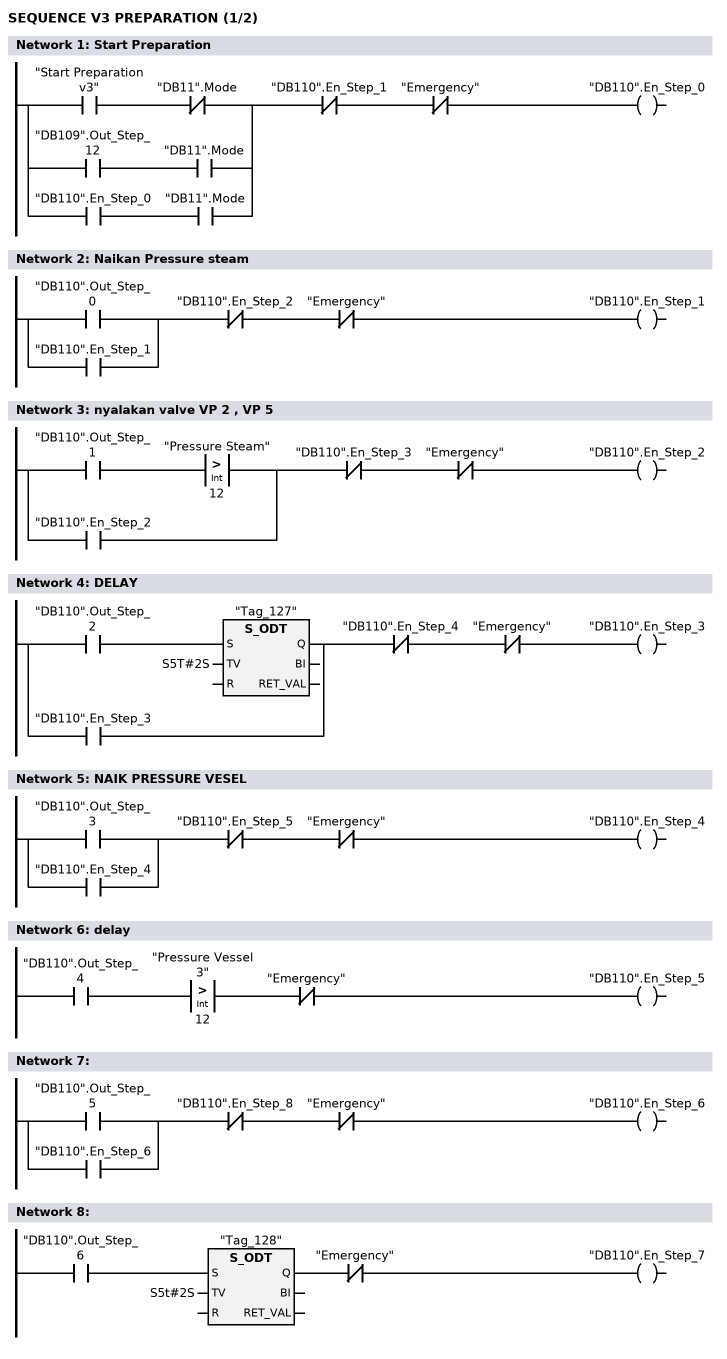
   RUNG wire#powerrail
      Contact( "Start Preparation v3" )
      I_Contact( "DB11".Mode )
      wire#w1
      I_Contact( "DB110".En_Step_1 )
      I_Contact( "Emergency" )
      Coil( "DB110".En_Step_0 )
   END_RUNG
   RUNG wire#powerrail
      Contact( "DB109".Out_Step_12 )
      Contact( "DB11".Mode )
   END_RUNG wire#w1
   RUNG wire#powerrail
      Contact( "DB110".En_Step_0 )
      Contact( "DB11".Mode )
   END_RUNG wire#w1
   // the same network as SCL:
   "DB110".En_Step_0 := (("Start Preparation v3" AND NOT "DB11".Mode) OR ("DB109".Out_Step_12 AND "DB11".Mode) OR ("DB110".En_Step_0 AND "DB11".Mode)) AND NOT "DB110".En_Step_1 AND NOT "Emergency";
END_REGION

REGION Network 2: Naikan Pressure steam
   RUNG wire#powerrail
      Contact( "DB110".Out_Step_0 )
      wire#w1
      I_Contact( "DB110".En_Step_2 )
      I_Contact( "Emergency" )
      Coil( "DB110".En_Step_1 )
   END_RUNG
   RUNG wire#powerrail
      Contact( "DB110".En_Step_1 )
   END_RUNG wire#w1
   // the same network as SCL:
   "DB110".En_Step_1 := ("DB110".Out_Step_0 OR "DB110".En_Step_1) AND NOT "DB110".En_Step_2 AND NOT "Emergency";
END_REGION

REGION Network 3: nyalakan valve VP 2 , VP 5
   RUNG wire#powerrail
      Contact( "DB110".Out_Step_1 )
      { S7_Templates := "SrcType := Int" } GT_Contact(in1 := "Pressure Steam", in2 := 12)
      wire#w1
      I_Contact( "DB110".En_Step_3 )
      I_Contact( "Emergency" )
      Coil( "DB110".En_Step_2 )
   END_RUNG
   RUNG wire#powerrail
      Contact( "DB110".En_Step_2 )
   END_RUNG wire#w1
   // the same network as SCL:
   "DB110".En_Step_2 := (("DB110".Out_Step_1 AND ("Pressure Steam" > 12)) OR "DB110".En_Step_2) AND NOT "DB110".En_Step_3 AND NOT "Emergency";
END_REGION

REGION Network 4: DELAY
   RUNG wire#powerrail
      Contact( "DB110".Out_Step_2 )
      S_ODT(T_NO := "Tag_127", TV := S5T#2S, R :=, BI =>, RET_VAL =>)
      wire#w1
      I_Contact( "DB110".En_Step_4 )
      I_Contact( "Emergency" )
      Coil( "DB110".En_Step_3 )
   END_RUNG
   RUNG wire#powerrail
      Contact( "DB110".En_Step_3 )
   END_RUNG wire#w1
   // the same network as SCL:
   #_s5time1 := S_ODT(T_NO := "Tag_127", S := "DB110".Out_Step_2, TV := S5T#2S, Q => #_w1);
   "DB110".En_Step_3 := (#_w1 OR "DB110".En_Step_3) AND NOT "DB110".En_Step_4 AND NOT "Emergency";
END_REGION

REGION Network 5: NAIK PRESSURE VESEL
   RUNG wire#powerrail
      Contact( "DB110".Out_Step_3 )
      wire#w1
      I_Contact( "DB110".En_Step_5 )
      I_Contact( "Emergency" )
      Coil( "DB110".En_Step_4 )
   END_RUNG
   RUNG wire#powerrail
      Contact( "DB110".En_Step_4 )
   END_RUNG wire#w1
   // the same network as SCL:
   "DB110".En_Step_4 := ("DB110".Out_Step_3 OR "DB110".En_Step_4) AND NOT "DB110".En_Step_5 AND NOT "Emergency";
END_REGION

REGION Network 6: delay
   RUNG wire#powerrail
      Contact( "DB110".Out_Step_4 )
      { S7_Templates := "SrcType := Int" } GT_Contact(in1 := "Pressure Vessel 3", in2 := 12)
      I_Contact( "Emergency" )
      Coil( "DB110".En_Step_5 )
   END_RUNG
   // the same network as SCL:
   "DB110".En_Step_5 := "DB110".Out_Step_4 AND ("Pressure Vessel 3" > 12) AND NOT "Emergency";
END_REGION

REGION Network 7
   RUNG wire#powerrail
      Contact( "DB110".Out_Step_5 )
      wire#w1
      I_Contact( "DB110".En_Step_8 )
      I_Contact( "Emergency" )
      Coil( "DB110".En_Step_6 )
   END_RUNG
   RUNG wire#powerrail
      Contact( "DB110".En_Step_6 )
   END_RUNG wire#w1
   // the same network as SCL:
   "DB110".En_Step_6 := ("DB110".Out_Step_5 OR "DB110".En_Step_6) AND NOT "DB110".En_Step_8 AND NOT "Emergency";
END_REGION

REGION Network 8
   RUNG wire#powerrail
      Contact( "DB110".Out_Step_6 )
      S_ODT(T_NO := "Tag_128", TV := S5t#2S, R :=, BI =>, RET_VAL =>)
      I_Contact( "Emergency" )
      Coil( "DB110".En_Step_7 )
   END_RUNG
   // the same network as SCL:
   #_s5time1 := S_ODT(T_NO := "Tag_128", S := "DB110".Out_Step_6, TV := S5t#2S, Q => #_w1);
   "DB110".En_Step_7 := #_w1 AND NOT "Emergency";
END_REGION

REGION Network 9: TURUNKAN PRESSURE
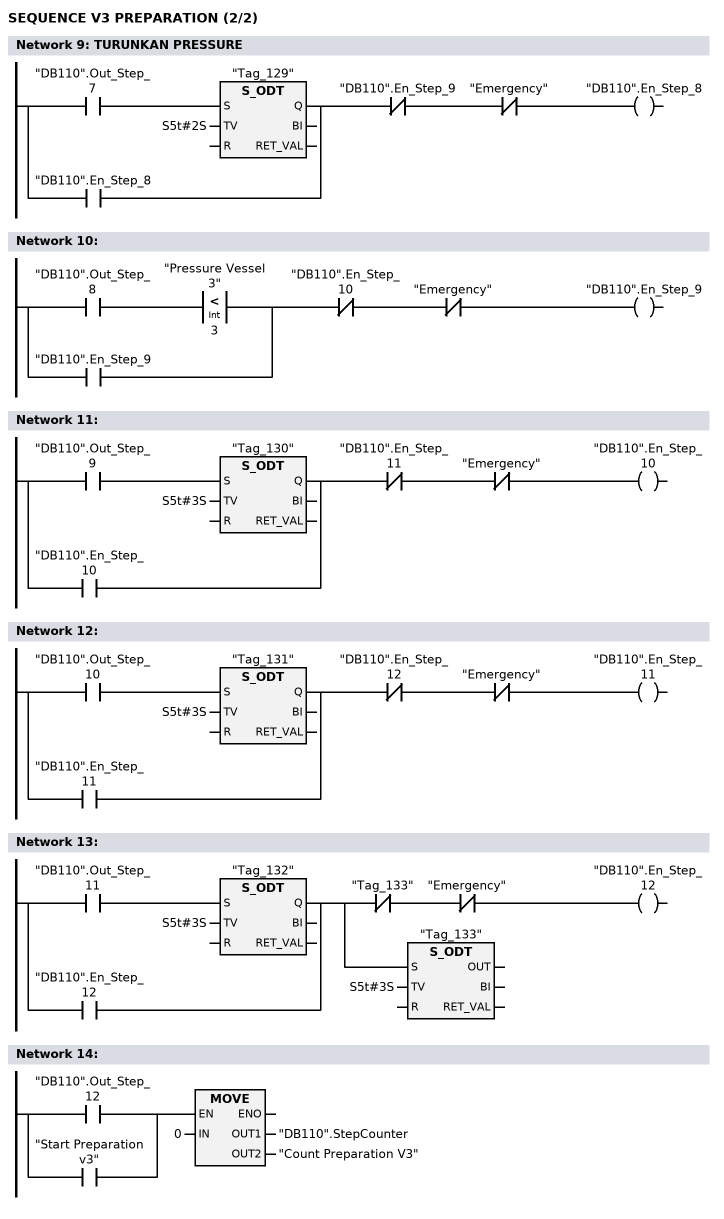
   RUNG wire#powerrail
      Contact( "DB110".Out_Step_7 )
      S_ODT(T_NO := "Tag_129", TV := S5t#2S, R :=, BI =>, RET_VAL =>)
      wire#w1
      I_Contact( "DB110".En_Step_9 )
      I_Contact( "Emergency" )
      Coil( "DB110".En_Step_8 )
   END_RUNG
   RUNG wire#powerrail
      Contact( "DB110".En_Step_8 )
   END_RUNG wire#w1
   // the same network as SCL:
   #_s5time1 := S_ODT(T_NO := "Tag_129", S := "DB110".Out_Step_7, TV := S5t#2S, Q => #_w1);
   "DB110".En_Step_8 := (#_w1 OR "DB110".En_Step_8) AND NOT "DB110".En_Step_9 AND NOT "Emergency";
END_REGION

REGION Network 10
   RUNG wire#powerrail
      Contact( "DB110".Out_Step_8 )
      { S7_Templates := "SrcType := Int" } LT_Contact(in1 := "Pressure Vessel 3", in2 := 3)
      wire#w1
      I_Contact( "DB110".En_Step_10 )
      I_Contact( "Emergency" )
      Coil( "DB110".En_Step_9 )
   END_RUNG
   RUNG wire#powerrail
      Contact( "DB110".En_Step_9 )
   END_RUNG wire#w1
   // the same network as SCL:
   "DB110".En_Step_9 := (("DB110".Out_Step_8 AND ("Pressure Vessel 3" < 3)) OR "DB110".En_Step_9) AND NOT "DB110".En_Step_10 AND NOT "Emergency";
END_REGION

REGION Network 11
   RUNG wire#powerrail
      Contact( "DB110".Out_Step_9 )
      S_ODT(T_NO := "Tag_130", TV := S5t#3S, R :=, BI =>, RET_VAL =>)
      wire#w1
      I_Contact( "DB110".En_Step_11 )
      I_Contact( "Emergency" )
      Coil( "DB110".En_Step_10 )
   END_RUNG
   RUNG wire#powerrail
      Contact( "DB110".En_Step_10 )
   END_RUNG wire#w1
   // the same network as SCL:
   #_s5time1 := S_ODT(T_NO := "Tag_130", S := "DB110".Out_Step_9, TV := S5t#3S, Q => #_w1);
   "DB110".En_Step_10 := (#_w1 OR "DB110".En_Step_10) AND NOT "DB110".En_Step_11 AND NOT "Emergency";
END_REGION

REGION Network 12
   RUNG wire#powerrail
      Contact( "DB110".Out_Step_10 )
      S_ODT(T_NO := "Tag_131", TV := S5t#3S, R :=, BI =>, RET_VAL =>)
      wire#w1
      I_Contact( "DB110".En_Step_12 )
      I_Contact( "Emergency" )
      Coil( "DB110".En_Step_11 )
   END_RUNG
   RUNG wire#powerrail
      Contact( "DB110".En_Step_11 )
   END_RUNG wire#w1
   // the same network as SCL:
   #_s5time1 := S_ODT(T_NO := "Tag_131", S := "DB110".Out_Step_10, TV := S5t#3S, Q => #_w1);
   "DB110".En_Step_11 := (#_w1 OR "DB110".En_Step_11) AND NOT "DB110".En_Step_12 AND NOT "Emergency";
END_REGION

REGION Network 13
   RUNG wire#powerrail
      Contact( "DB110".Out_Step_11 )
      S_ODT(T_NO := "Tag_132", TV := S5t#3S, R :=, BI =>, RET_VAL =>)
      wire#w1
      I_Contact( "Tag_133" )
      I_Contact( "Emergency" )
      Coil( "DB110".En_Step_12 )
   END_RUNG
   RUNG wire#powerrail
      Contact( "DB110".En_Step_12 )
   END_RUNG wire#w1
   RUNG wire#w1
      S_ODT(T_NO := "Tag_133", TV := S5t#3S, R :=, BI =>, RET_VAL =>)
   END_RUNG
   // the same network as SCL:
   #_s5time1 := S_ODT(T_NO := "Tag_132", S := "DB110".Out_Step_11, TV := S5t#3S, Q => #_w1);
   #_w2 := #_w1 OR "DB110".En_Step_12;
   "DB110".En_Step_12 := #_w2 AND NOT "Tag_133" AND NOT "Emergency";
   #_s5time2 := S_ODT(T_NO := "Tag_133", S := #_w2, TV := S5t#3S);
END_REGION

REGION Network 14
   RUNG wire#powerrail
      Contact( "DB110".Out_Step_12 )
      wire#w1
      Move(in := 0, out1 => "DB110".StepCounter, out2 => "Count Preparation V3")
   END_RUNG
   RUNG wire#powerrail
      Contact( "Start Preparation v3" )
   END_RUNG wire#w1
   // the same network as SCL:
   IF "DB110".Out_Step_12 OR "Start Preparation v3" THEN
       "DB110".StepCounter := 0;
       "Count Preparation V3" := 0;
   END_IF;
END_REGION
END_FUNCTION

FUNCTION "VESSEL 3 PREPARATION" : Void   // FC26, LAD
{ S7_Optimized_Access := 'TRUE' }
VERSION : 0.1
   VAR_TEMP   // added for the SCL form of the ladder/FBD networks
      _w1 : Bool;
      _w2 : Bool;
      _w3 : Bool;
      _w4 : Bool;
   END_VAR
BEGIN

REGION Network 1: NAIKAN PRESSURE STEAM
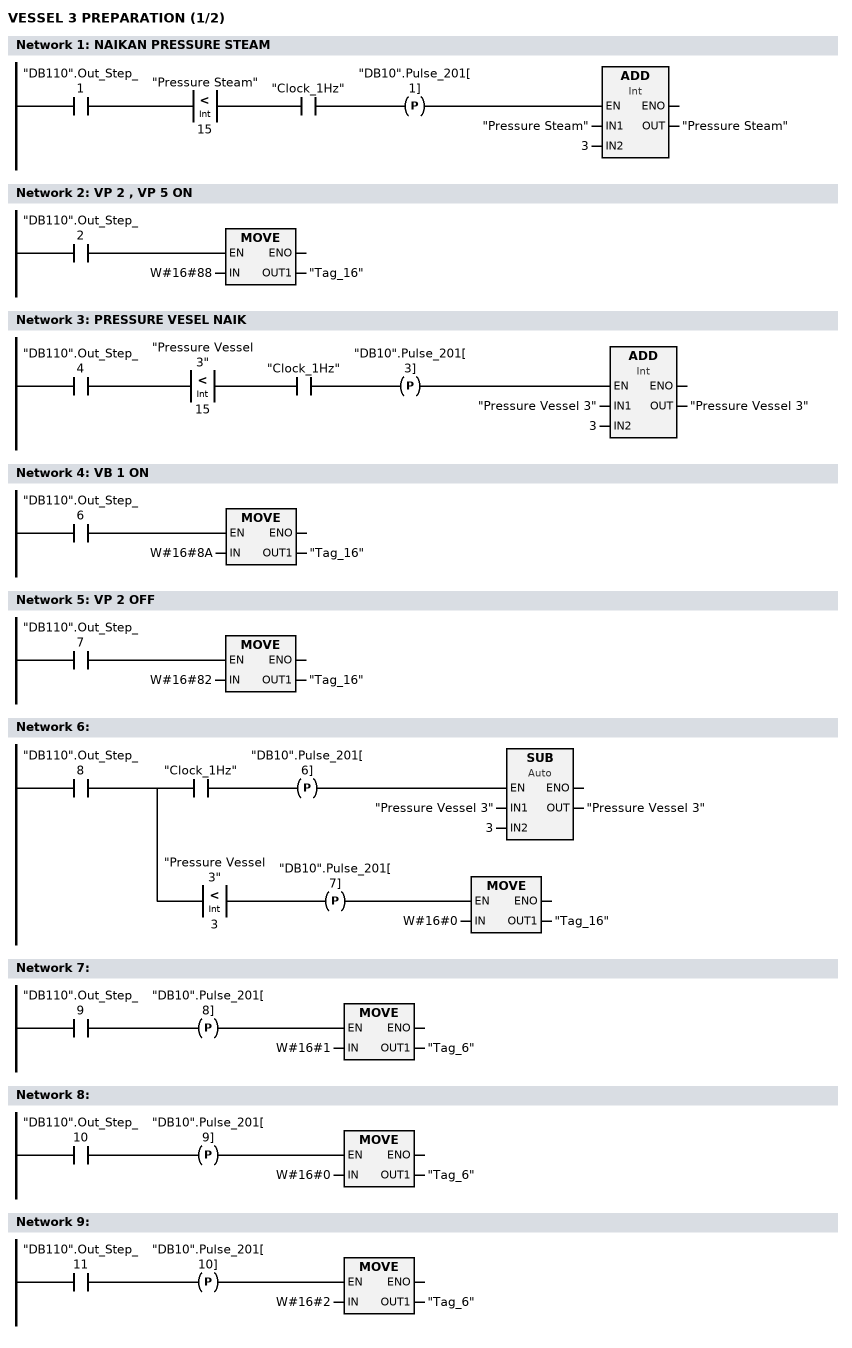
   RUNG wire#powerrail
      Contact( "DB110".Out_Step_1 )
      { S7_Templates := "SrcType := Int" } LT_Contact(in1 := "Pressure Steam", in2 := 15)
      Contact( "Clock_1Hz" )
      P_Trig( "DB10".Pulse_201[1] )
      { S7_Templates := "SrcType := Int" } Add(in1 := "Pressure Steam", in2 := 3, out => "Pressure Steam")
   END_RUNG
   // the same network as SCL:
   #_w1 := "DB110".Out_Step_1 AND ("Pressure Steam" < 15) AND "Clock_1Hz";
   #_w2 := #_w1 AND NOT "DB10".Pulse_201[1];   // rising edge
   "DB10".Pulse_201[1] := #_w1;
   IF #_w2 THEN "Pressure Steam" := "Pressure Steam" + 3; END_IF;
END_REGION

REGION Network 2: VP 2 , VP 5 ON
   RUNG wire#powerrail
      Contact( "DB110".Out_Step_2 )
      Move(in := W#16#88, out1 => "Tag_16")
   END_RUNG
   // the same network as SCL:
   IF "DB110".Out_Step_2 THEN "Tag_16" := W#16#88; END_IF;
END_REGION

REGION Network 3: PRESSURE VESEL NAIK
   RUNG wire#powerrail
      Contact( "DB110".Out_Step_4 )
      { S7_Templates := "SrcType := Int" } LT_Contact(in1 := "Pressure Vessel 3", in2 := 15)
      Contact( "Clock_1Hz" )
      P_Trig( "DB10".Pulse_201[3] )
      { S7_Templates := "SrcType := Int" } Add(in1 := "Pressure Vessel 3", in2 := 3, out => "Pressure Vessel 3")
   END_RUNG
   // the same network as SCL:
   #_w1 := "DB110".Out_Step_4 AND ("Pressure Vessel 3" < 15) AND "Clock_1Hz";
   #_w2 := #_w1 AND NOT "DB10".Pulse_201[3];   // rising edge
   "DB10".Pulse_201[3] := #_w1;
   IF #_w2 THEN "Pressure Vessel 3" := "Pressure Vessel 3" + 3; END_IF;
END_REGION

REGION Network 4: VB 1 ON
   RUNG wire#powerrail
      Contact( "DB110".Out_Step_6 )
      Move(in := W#16#8A, out1 => "Tag_16")
   END_RUNG
   // the same network as SCL:
   IF "DB110".Out_Step_6 THEN "Tag_16" := W#16#8A; END_IF;
END_REGION

REGION Network 5: VP 2 OFF
   RUNG wire#powerrail
      Contact( "DB110".Out_Step_7 )
      Move(in := W#16#82, out1 => "Tag_16")
   END_RUNG
   // the same network as SCL:
   IF "DB110".Out_Step_7 THEN "Tag_16" := W#16#82; END_IF;
END_REGION

REGION Network 6
   RUNG wire#powerrail
      Contact( "DB110".Out_Step_8 )
      wire#w1
      Contact( "Clock_1Hz" )
      P_Trig( "DB10".Pulse_201[6] )
      Sub(in1 := "Pressure Vessel 3", in2 := 3, out => "Pressure Vessel 3")
   END_RUNG
   RUNG wire#w1
      { S7_Templates := "SrcType := Int" } LT_Contact(in1 := "Pressure Vessel 3", in2 := 3)
      P_Trig( "DB10".Pulse_201[7] )
      Move(in := W#16#0, out1 => "Tag_16")
   END_RUNG
   // the same network as SCL:
   #_w1 := "DB110".Out_Step_8 AND "Clock_1Hz";
   #_w2 := #_w1 AND NOT "DB10".Pulse_201[6];   // rising edge
   "DB10".Pulse_201[6] := #_w1;
   IF #_w2 THEN "Pressure Vessel 3" := "Pressure Vessel 3" - 3; END_IF;
   #_w3 := "DB110".Out_Step_8 AND ("Pressure Vessel 3" < 3);
   #_w4 := #_w3 AND NOT "DB10".Pulse_201[7];   // rising edge
   "DB10".Pulse_201[7] := #_w3;
   IF #_w4 THEN "Tag_16" := W#16#0; END_IF;
END_REGION

REGION Network 7
   RUNG wire#powerrail
      Contact( "DB110".Out_Step_9 )
      P_Trig( "DB10".Pulse_201[8] )
      Move(in := W#16#1, out1 => "Tag_6")
   END_RUNG
   // the same network as SCL:
   #_w1 := "DB110".Out_Step_9 AND NOT "DB10".Pulse_201[8];   // rising edge
   "DB10".Pulse_201[8] := "DB110".Out_Step_9;
   IF #_w1 THEN "Tag_6" := W#16#1; END_IF;
END_REGION

REGION Network 8
   RUNG wire#powerrail
      Contact( "DB110".Out_Step_10 )
      P_Trig( "DB10".Pulse_201[9] )
      Move(in := W#16#0, out1 => "Tag_6")
   END_RUNG
   // the same network as SCL:
   #_w1 := "DB110".Out_Step_10 AND NOT "DB10".Pulse_201[9];   // rising edge
   "DB10".Pulse_201[9] := "DB110".Out_Step_10;
   IF #_w1 THEN "Tag_6" := W#16#0; END_IF;
END_REGION

REGION Network 9
   RUNG wire#powerrail
      Contact( "DB110".Out_Step_11 )
      P_Trig( "DB10".Pulse_201[10] )
      Move(in := W#16#2, out1 => "Tag_6")
   END_RUNG
   // the same network as SCL:
   #_w1 := "DB110".Out_Step_11 AND NOT "DB10".Pulse_201[10];   // rising edge
   "DB10".Pulse_201[10] := "DB110".Out_Step_11;
   IF #_w1 THEN "Tag_6" := W#16#2; END_IF;
END_REGION

REGION Network 10
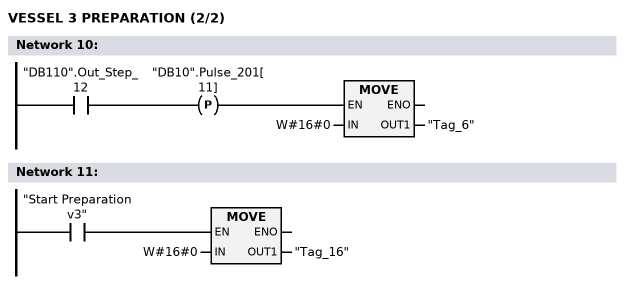
   RUNG wire#powerrail
      Contact( "DB110".Out_Step_12 )
      P_Trig( "DB10".Pulse_201[11] )
      Move(in := W#16#0, out1 => "Tag_6")
   END_RUNG
   // the same network as SCL:
   #_w1 := "DB110".Out_Step_12 AND NOT "DB10".Pulse_201[11];   // rising edge
   "DB10".Pulse_201[11] := "DB110".Out_Step_12;
   IF #_w1 THEN "Tag_6" := W#16#0; END_IF;
END_REGION

REGION Network 11
   RUNG wire#powerrail
      Contact( "Start Preparation v3" )
      Move(in := W#16#0, out1 => "Tag_16")
   END_RUNG
   // the same network as SCL:
   IF "Start Preparation v3" THEN "Tag_16" := W#16#0; END_IF;
END_REGION
END_FUNCTION

FUNCTION "SEQUENCE V4 PREPARATION" : Void   // FC27, LAD
{ S7_Optimized_Access := 'TRUE' }
VERSION : 0.1
   VAR_TEMP   // added for the SCL form of the ladder/FBD networks
      _w1 : Bool;
      _s5time1 : S5Time;
      _w2 : Bool;
      _s5time2 : S5Time;
   END_VAR
BEGIN

REGION Network 1: Start Preparation
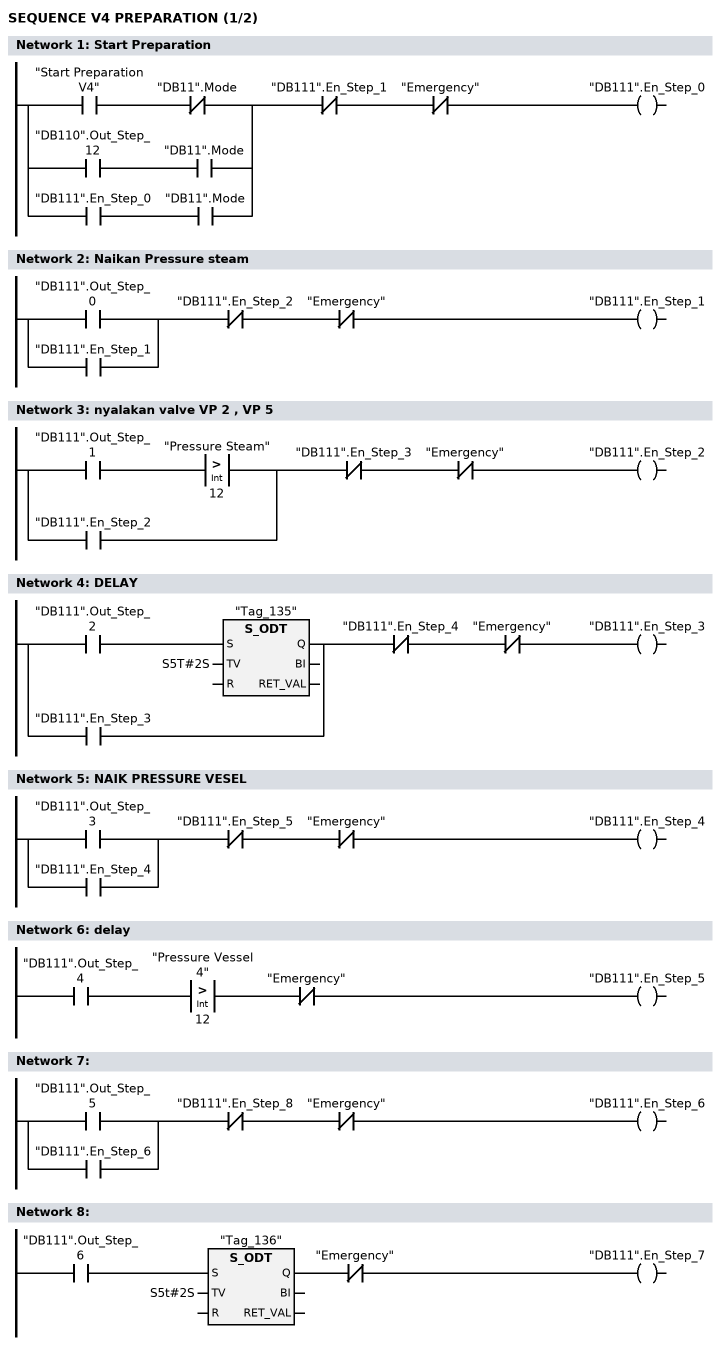
   RUNG wire#powerrail
      Contact( "Start Preparation V4" )
      I_Contact( "DB11".Mode )
      wire#w1
      I_Contact( "DB111".En_Step_1 )
      I_Contact( "Emergency" )
      Coil( "DB111".En_Step_0 )
   END_RUNG
   RUNG wire#powerrail
      Contact( "DB110".Out_Step_12 )
      Contact( "DB11".Mode )
   END_RUNG wire#w1
   RUNG wire#powerrail
      Contact( "DB111".En_Step_0 )
      Contact( "DB11".Mode )
   END_RUNG wire#w1
   // the same network as SCL:
   "DB111".En_Step_0 := (("Start Preparation V4" AND NOT "DB11".Mode) OR ("DB110".Out_Step_12 AND "DB11".Mode) OR ("DB111".En_Step_0 AND "DB11".Mode)) AND NOT "DB111".En_Step_1 AND NOT "Emergency";
END_REGION

REGION Network 2: Naikan Pressure steam
   RUNG wire#powerrail
      Contact( "DB111".Out_Step_0 )
      wire#w1
      I_Contact( "DB111".En_Step_2 )
      I_Contact( "Emergency" )
      Coil( "DB111".En_Step_1 )
   END_RUNG
   RUNG wire#powerrail
      Contact( "DB111".En_Step_1 )
   END_RUNG wire#w1
   // the same network as SCL:
   "DB111".En_Step_1 := ("DB111".Out_Step_0 OR "DB111".En_Step_1) AND NOT "DB111".En_Step_2 AND NOT "Emergency";
END_REGION

REGION Network 3: nyalakan valve VP 2 , VP 5
   RUNG wire#powerrail
      Contact( "DB111".Out_Step_1 )
      { S7_Templates := "SrcType := Int" } GT_Contact(in1 := "Pressure Steam", in2 := 12)
      wire#w1
      I_Contact( "DB111".En_Step_3 )
      I_Contact( "Emergency" )
      Coil( "DB111".En_Step_2 )
   END_RUNG
   RUNG wire#powerrail
      Contact( "DB111".En_Step_2 )
   END_RUNG wire#w1
   // the same network as SCL:
   "DB111".En_Step_2 := (("DB111".Out_Step_1 AND ("Pressure Steam" > 12)) OR "DB111".En_Step_2) AND NOT "DB111".En_Step_3 AND NOT "Emergency";
END_REGION

REGION Network 4: DELAY
   RUNG wire#powerrail
      Contact( "DB111".Out_Step_2 )
      S_ODT(T_NO := "Tag_135", TV := S5T#2S, R :=, BI =>, RET_VAL =>)
      wire#w1
      I_Contact( "DB111".En_Step_4 )
      I_Contact( "Emergency" )
      Coil( "DB111".En_Step_3 )
   END_RUNG
   RUNG wire#powerrail
      Contact( "DB111".En_Step_3 )
   END_RUNG wire#w1
   // the same network as SCL:
   #_s5time1 := S_ODT(T_NO := "Tag_135", S := "DB111".Out_Step_2, TV := S5T#2S, Q => #_w1);
   "DB111".En_Step_3 := (#_w1 OR "DB111".En_Step_3) AND NOT "DB111".En_Step_4 AND NOT "Emergency";
END_REGION

REGION Network 5: NAIK PRESSURE VESEL
   RUNG wire#powerrail
      Contact( "DB111".Out_Step_3 )
      wire#w1
      I_Contact( "DB111".En_Step_5 )
      I_Contact( "Emergency" )
      Coil( "DB111".En_Step_4 )
   END_RUNG
   RUNG wire#powerrail
      Contact( "DB111".En_Step_4 )
   END_RUNG wire#w1
   // the same network as SCL:
   "DB111".En_Step_4 := ("DB111".Out_Step_3 OR "DB111".En_Step_4) AND NOT "DB111".En_Step_5 AND NOT "Emergency";
END_REGION

REGION Network 6: delay
   RUNG wire#powerrail
      Contact( "DB111".Out_Step_4 )
      { S7_Templates := "SrcType := Int" } GT_Contact(in1 := "Pressure Vessel 4", in2 := 12)
      I_Contact( "Emergency" )
      Coil( "DB111".En_Step_5 )
   END_RUNG
   // the same network as SCL:
   "DB111".En_Step_5 := "DB111".Out_Step_4 AND ("Pressure Vessel 4" > 12) AND NOT "Emergency";
END_REGION

REGION Network 7
   RUNG wire#powerrail
      Contact( "DB111".Out_Step_5 )
      wire#w1
      I_Contact( "DB111".En_Step_8 )
      I_Contact( "Emergency" )
      Coil( "DB111".En_Step_6 )
   END_RUNG
   RUNG wire#powerrail
      Contact( "DB111".En_Step_6 )
   END_RUNG wire#w1
   // the same network as SCL:
   "DB111".En_Step_6 := ("DB111".Out_Step_5 OR "DB111".En_Step_6) AND NOT "DB111".En_Step_8 AND NOT "Emergency";
END_REGION

REGION Network 8
   RUNG wire#powerrail
      Contact( "DB111".Out_Step_6 )
      S_ODT(T_NO := "Tag_136", TV := S5t#2S, R :=, BI =>, RET_VAL =>)
      I_Contact( "Emergency" )
      Coil( "DB111".En_Step_7 )
   END_RUNG
   // the same network as SCL:
   #_s5time1 := S_ODT(T_NO := "Tag_136", S := "DB111".Out_Step_6, TV := S5t#2S, Q => #_w1);
   "DB111".En_Step_7 := #_w1 AND NOT "Emergency";
END_REGION

REGION Network 9: TURUNKAN PRESSURE
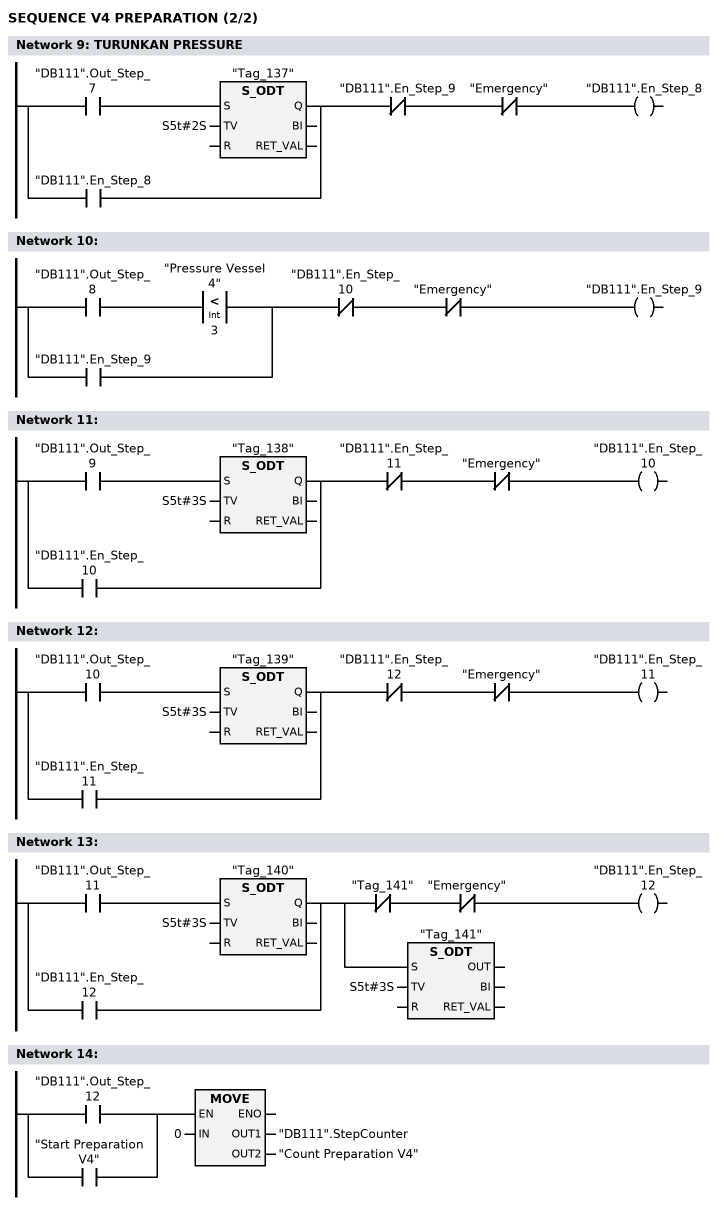
   RUNG wire#powerrail
      Contact( "DB111".Out_Step_7 )
      S_ODT(T_NO := "Tag_137", TV := S5t#2S, R :=, BI =>, RET_VAL =>)
      wire#w1
      I_Contact( "DB111".En_Step_9 )
      I_Contact( "Emergency" )
      Coil( "DB111".En_Step_8 )
   END_RUNG
   RUNG wire#powerrail
      Contact( "DB111".En_Step_8 )
   END_RUNG wire#w1
   // the same network as SCL:
   #_s5time1 := S_ODT(T_NO := "Tag_137", S := "DB111".Out_Step_7, TV := S5t#2S, Q => #_w1);
   "DB111".En_Step_8 := (#_w1 OR "DB111".En_Step_8) AND NOT "DB111".En_Step_9 AND NOT "Emergency";
END_REGION

REGION Network 10
   RUNG wire#powerrail
      Contact( "DB111".Out_Step_8 )
      { S7_Templates := "SrcType := Int" } LT_Contact(in1 := "Pressure Vessel 4", in2 := 3)
      wire#w1
      I_Contact( "DB111".En_Step_10 )
      I_Contact( "Emergency" )
      Coil( "DB111".En_Step_9 )
   END_RUNG
   RUNG wire#powerrail
      Contact( "DB111".En_Step_9 )
   END_RUNG wire#w1
   // the same network as SCL:
   "DB111".En_Step_9 := (("DB111".Out_Step_8 AND ("Pressure Vessel 4" < 3)) OR "DB111".En_Step_9) AND NOT "DB111".En_Step_10 AND NOT "Emergency";
END_REGION

REGION Network 11
   RUNG wire#powerrail
      Contact( "DB111".Out_Step_9 )
      S_ODT(T_NO := "Tag_138", TV := S5t#3S, R :=, BI =>, RET_VAL =>)
      wire#w1
      I_Contact( "DB111".En_Step_11 )
      I_Contact( "Emergency" )
      Coil( "DB111".En_Step_10 )
   END_RUNG
   RUNG wire#powerrail
      Contact( "DB111".En_Step_10 )
   END_RUNG wire#w1
   // the same network as SCL:
   #_s5time1 := S_ODT(T_NO := "Tag_138", S := "DB111".Out_Step_9, TV := S5t#3S, Q => #_w1);
   "DB111".En_Step_10 := (#_w1 OR "DB111".En_Step_10) AND NOT "DB111".En_Step_11 AND NOT "Emergency";
END_REGION

REGION Network 12
   RUNG wire#powerrail
      Contact( "DB111".Out_Step_10 )
      S_ODT(T_NO := "Tag_139", TV := S5t#3S, R :=, BI =>, RET_VAL =>)
      wire#w1
      I_Contact( "DB111".En_Step_12 )
      I_Contact( "Emergency" )
      Coil( "DB111".En_Step_11 )
   END_RUNG
   RUNG wire#powerrail
      Contact( "DB111".En_Step_11 )
   END_RUNG wire#w1
   // the same network as SCL:
   #_s5time1 := S_ODT(T_NO := "Tag_139", S := "DB111".Out_Step_10, TV := S5t#3S, Q => #_w1);
   "DB111".En_Step_11 := (#_w1 OR "DB111".En_Step_11) AND NOT "DB111".En_Step_12 AND NOT "Emergency";
END_REGION

REGION Network 13
   RUNG wire#powerrail
      Contact( "DB111".Out_Step_11 )
      S_ODT(T_NO := "Tag_140", TV := S5t#3S, R :=, BI =>, RET_VAL =>)
      wire#w1
      I_Contact( "Tag_141" )
      I_Contact( "Emergency" )
      Coil( "DB111".En_Step_12 )
   END_RUNG
   RUNG wire#powerrail
      Contact( "DB111".En_Step_12 )
   END_RUNG wire#w1
   RUNG wire#w1
      S_ODT(T_NO := "Tag_141", TV := S5t#3S, R :=, BI =>, RET_VAL =>)
   END_RUNG
   // the same network as SCL:
   #_s5time1 := S_ODT(T_NO := "Tag_140", S := "DB111".Out_Step_11, TV := S5t#3S, Q => #_w1);
   #_w2 := #_w1 OR "DB111".En_Step_12;
   "DB111".En_Step_12 := #_w2 AND NOT "Tag_141" AND NOT "Emergency";
   #_s5time2 := S_ODT(T_NO := "Tag_141", S := #_w2, TV := S5t#3S);
END_REGION

REGION Network 14
   RUNG wire#powerrail
      Contact( "DB111".Out_Step_12 )
      wire#w1
      Move(in := 0, out1 => "DB111".StepCounter, out2 => "Count Preparation V4")
   END_RUNG
   RUNG wire#powerrail
      Contact( "Start Preparation V4" )
   END_RUNG wire#w1
   // the same network as SCL:
   IF "DB111".Out_Step_12 OR "Start Preparation V4" THEN
       "DB111".StepCounter := 0;
       "Count Preparation V4" := 0;
   END_IF;
END_REGION
END_FUNCTION

FUNCTION "VESSEL 4 PREPARATION" : Void   // FC28, LAD
{ S7_Optimized_Access := 'TRUE' }
VERSION : 0.1
   VAR_TEMP   // added for the SCL form of the ladder/FBD networks
      _w1 : Bool;
      _w2 : Bool;
      _w3 : Bool;
      _w4 : Bool;
   END_VAR
BEGIN

REGION Network 1: NAIKAN PRESSURE STEAM
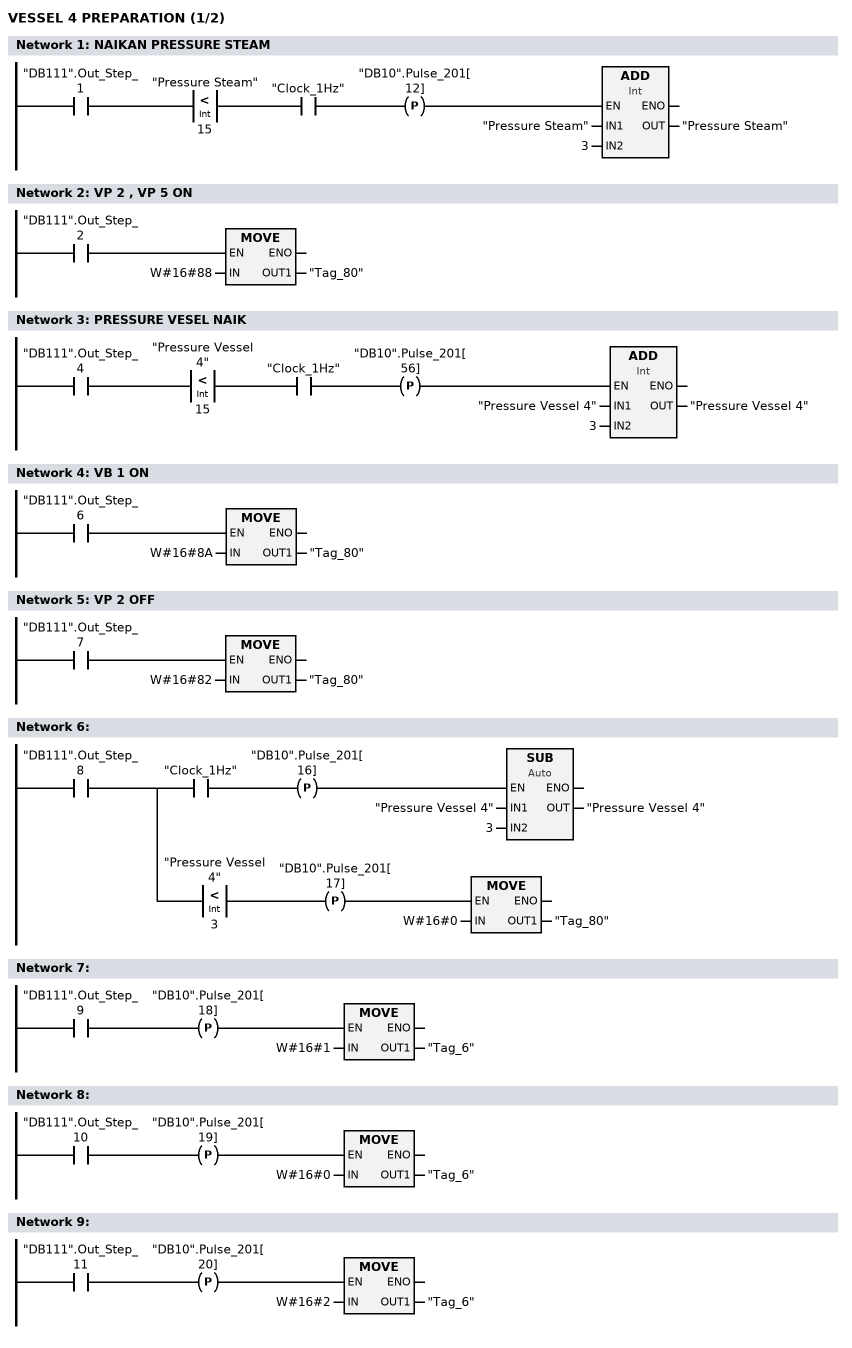
   RUNG wire#powerrail
      Contact( "DB111".Out_Step_1 )
      { S7_Templates := "SrcType := Int" } LT_Contact(in1 := "Pressure Steam", in2 := 15)
      Contact( "Clock_1Hz" )
      P_Trig( "DB10".Pulse_201[12] )
      { S7_Templates := "SrcType := Int" } Add(in1 := "Pressure Steam", in2 := 3, out => "Pressure Steam")
   END_RUNG
   // the same network as SCL:
   #_w1 := "DB111".Out_Step_1 AND ("Pressure Steam" < 15) AND "Clock_1Hz";
   #_w2 := #_w1 AND NOT "DB10".Pulse_201[12];   // rising edge
   "DB10".Pulse_201[12] := #_w1;
   IF #_w2 THEN "Pressure Steam" := "Pressure Steam" + 3; END_IF;
END_REGION

REGION Network 2: VP 2 , VP 5 ON
   RUNG wire#powerrail
      Contact( "DB111".Out_Step_2 )
      Move(in := W#16#88, out1 => "Tag_80")
   END_RUNG
   // the same network as SCL:
   IF "DB111".Out_Step_2 THEN "Tag_80" := W#16#88; END_IF;
END_REGION

REGION Network 3: PRESSURE VESEL NAIK
   RUNG wire#powerrail
      Contact( "DB111".Out_Step_4 )
      { S7_Templates := "SrcType := Int" } LT_Contact(in1 := "Pressure Vessel 4", in2 := 15)
      Contact( "Clock_1Hz" )
      P_Trig( "DB10".Pulse_201[56] )
      { S7_Templates := "SrcType := Int" } Add(in1 := "Pressure Vessel 4", in2 := 3, out => "Pressure Vessel 4")
   END_RUNG
   // the same network as SCL:
   #_w1 := "DB111".Out_Step_4 AND ("Pressure Vessel 4" < 15) AND "Clock_1Hz";
   #_w2 := #_w1 AND NOT "DB10".Pulse_201[56];   // rising edge
   "DB10".Pulse_201[56] := #_w1;
   IF #_w2 THEN "Pressure Vessel 4" := "Pressure Vessel 4" + 3; END_IF;
END_REGION

REGION Network 4: VB 1 ON
   RUNG wire#powerrail
      Contact( "DB111".Out_Step_6 )
      Move(in := W#16#8A, out1 => "Tag_80")
   END_RUNG
   // the same network as SCL:
   IF "DB111".Out_Step_6 THEN "Tag_80" := W#16#8A; END_IF;
END_REGION

REGION Network 5: VP 2 OFF
   RUNG wire#powerrail
      Contact( "DB111".Out_Step_7 )
      Move(in := W#16#82, out1 => "Tag_80")
   END_RUNG
   // the same network as SCL:
   IF "DB111".Out_Step_7 THEN "Tag_80" := W#16#82; END_IF;
END_REGION

REGION Network 6
   RUNG wire#powerrail
      Contact( "DB111".Out_Step_8 )
      wire#w1
      Contact( "Clock_1Hz" )
      P_Trig( "DB10".Pulse_201[16] )
      Sub(in1 := "Pressure Vessel 4", in2 := 3, out => "Pressure Vessel 4")
   END_RUNG
   RUNG wire#w1
      { S7_Templates := "SrcType := Int" } LT_Contact(in1 := "Pressure Vessel 4", in2 := 3)
      P_Trig( "DB10".Pulse_201[17] )
      Move(in := W#16#0, out1 => "Tag_80")
   END_RUNG
   // the same network as SCL:
   #_w1 := "DB111".Out_Step_8 AND "Clock_1Hz";
   #_w2 := #_w1 AND NOT "DB10".Pulse_201[16];   // rising edge
   "DB10".Pulse_201[16] := #_w1;
   IF #_w2 THEN "Pressure Vessel 4" := "Pressure Vessel 4" - 3; END_IF;
   #_w3 := "DB111".Out_Step_8 AND ("Pressure Vessel 4" < 3);
   #_w4 := #_w3 AND NOT "DB10".Pulse_201[17];   // rising edge
   "DB10".Pulse_201[17] := #_w3;
   IF #_w4 THEN "Tag_80" := W#16#0; END_IF;
END_REGION

REGION Network 7
   RUNG wire#powerrail
      Contact( "DB111".Out_Step_9 )
      P_Trig( "DB10".Pulse_201[18] )
      Move(in := W#16#1, out1 => "Tag_6")
   END_RUNG
   // the same network as SCL:
   #_w1 := "DB111".Out_Step_9 AND NOT "DB10".Pulse_201[18];   // rising edge
   "DB10".Pulse_201[18] := "DB111".Out_Step_9;
   IF #_w1 THEN "Tag_6" := W#16#1; END_IF;
END_REGION

REGION Network 8
   RUNG wire#powerrail
      Contact( "DB111".Out_Step_10 )
      P_Trig( "DB10".Pulse_201[19] )
      Move(in := W#16#0, out1 => "Tag_6")
   END_RUNG
   // the same network as SCL:
   #_w1 := "DB111".Out_Step_10 AND NOT "DB10".Pulse_201[19];   // rising edge
   "DB10".Pulse_201[19] := "DB111".Out_Step_10;
   IF #_w1 THEN "Tag_6" := W#16#0; END_IF;
END_REGION

REGION Network 9
   RUNG wire#powerrail
      Contact( "DB111".Out_Step_11 )
      P_Trig( "DB10".Pulse_201[20] )
      Move(in := W#16#2, out1 => "Tag_6")
   END_RUNG
   // the same network as SCL:
   #_w1 := "DB111".Out_Step_11 AND NOT "DB10".Pulse_201[20];   // rising edge
   "DB10".Pulse_201[20] := "DB111".Out_Step_11;
   IF #_w1 THEN "Tag_6" := W#16#2; END_IF;
END_REGION

REGION Network 10
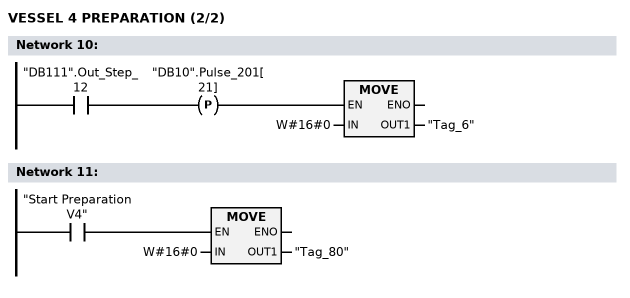
   RUNG wire#powerrail
      Contact( "DB111".Out_Step_12 )
      P_Trig( "DB10".Pulse_201[21] )
      Move(in := W#16#0, out1 => "Tag_6")
   END_RUNG
   // the same network as SCL:
   #_w1 := "DB111".Out_Step_12 AND NOT "DB10".Pulse_201[21];   // rising edge
   "DB10".Pulse_201[21] := "DB111".Out_Step_12;
   IF #_w1 THEN "Tag_6" := W#16#0; END_IF;
END_REGION

REGION Network 11
   RUNG wire#powerrail
      Contact( "Start Preparation V4" )
      Move(in := W#16#0, out1 => "Tag_80")
   END_RUNG
   // the same network as SCL:
   IF "Start Preparation V4" THEN "Tag_80" := W#16#0; END_IF;
END_REGION
END_FUNCTION

FUNCTION "SEQUENCE V5 PREPARATION" : Void   // FC29, LAD
{ S7_Optimized_Access := 'TRUE' }
VERSION : 0.1
   VAR_TEMP   // added for the SCL form of the ladder/FBD networks
      _w1 : Bool;
      _s5time1 : S5Time;
      _w2 : Bool;
      _s5time2 : S5Time;
   END_VAR
BEGIN

REGION Network 1: Start Preparation
